screen "Inert Gas Generator Plant" 1280x800, template "Template"
   GraphicView "Graphic view_52" at 522,118 size 43x67; Picture "Graphic_72"
   GraphicView "Graphic view_49" at 715,199 size 43x67; Picture "Graphic_72"
   GraphicView "Graphic view_12" at 522,199 size 43x67; Picture "Graphic_72"
   GraphicView "Graphic view_55" at 522,416 size 43x67; Picture "Graphic_72"
   GraphicView "Graphic view_56" at 650,416 size 43x67; Picture "Graphic_72"
   GraphicView "Graphic view_57" at 522,311 size 43x67; Picture "Graphic_72"
   GraphicView "Graphic view_61" at 527,525 size 32x54; Picture "Graphic_72"
   TextField "Text field_97" at 742,724 size 131x20; Text 'IGG Gas Pressure'
   TextField "Text field_98" at 866,724 size 147x20; Text 'Atom. Air Pressure'
   TextField "Text field_47" at 251,73 size 69x18; Text 'Full Auto'
      Visibility <- "82_To_HMI_CRNT_MODE_IGG"
   TextField "Text field_1" at 251,74 size 55x18; Text 'Manual'
      Visibility <- "82_To_HMI_CRNT_MODE_IGG"
   TextField "Text field_4" at 252,74 size 103x18; Text 'Undetermined'
      Visibility <- "82_To_HMI_CRNT_MODE_IGG"
   TextField "Text field_57" at 252,74 size 36x18; Text 'FAT'
      Visibility <- "82_To_HMI_CRNT_MODE_IGG"
   TextField "Text field_42" at 434,121 size 70x22; Text 'No Flow'
   TextField "Text field_43" at 434,121 size 70x22; Text '- Flow -'
      Visibility <- "10 DI_DATA_FS123"
      Appearance <- "10 DI_DATA_FS123"
   GraphicView "Logo" at 1,1 size 219x60; Picture "Logo of IGG HMI"
   Group "Group_8" at 743,722 size 397x61
   Button "Button_1" at 902,751 size 66x25; TextOn 'Enabled'; TextOff 'Text'
   IOField "I/O field_29" at 898,751 size 70x25; Authorization "Commissioning"; FormatPattern 99.99; Unit  bar
      ProcessValue <- "1111_PID_CV111_Setpoint"
   Group "Group" at 742,724 size 271x20
   IOField "I/O field_10" at 956,109 size 54x22; FormatPattern 999; Unit %
      ProcessValue <- "12_AI_Data_CV403_SCALED"
   IOField "I/O field_15" at 956,95 size 54x22; FormatPattern 999; Unit %
      ProcessValue <- "16_AQ_Data_CV403_CNTRL"
   GraphicView "Graphic view_5" at 1149,212 size 128x29; Picture "Graphic_82"
   GraphicView "Graphic view_91" at 22,264 size 113x127; Picture "Graphic_246"
   GraphicIOField "Graphic I/O field_5" at 14,257 size 129x139; PictureList "New IA Compressor"
      ProcessValue <- "82_To_HMI_IA Compressor Animation"
      Visibility <- "68_Sys_Status_Data_IA_PRES_IN_RNG(1)"
   GraphicView "Graphic view_93" at 147,261 size 48x132; Picture "Graphic_248"
   TextField "Text field_58" at 41,731 size 135x20; Text 'Fuel Pump System'
      Appearance <- "68_Sys_Status_Data_FUEL_PRES_IN_RNG"
   TextField "Text field_89" at 1115,538 size 54x22; Text 'Text'
   Button "HmiScreenItemData_1" at 1,50 size 150x43; TextOn 'Back'; TextOff 'Main Index'
      on Release: ActivateScreen("02 Main Index", 0)
   GraphicView "Graphic view_20" at 336,126 size 900x542; Picture "IGG_5"
   GraphicView "Graphic view_41" at 815,266 size 13x60; Picture "Graphic_57"
   GraphicView "Graphic view_11" at 296,251 size 377x12; Picture "Graphic_20"
   GraphicView "Graphic view_40" at 806,251 size 21x20; Picture "Graphic_41"
   GraphicView "Graphic view_42" at 296,468 size 278x12; Picture "Graphic_20"
   GraphicView "Graphic view_43" at 696,458 size 19x21; Picture "Graphic_40"
   GraphicView "Graphic view_44" at 294,251 size 20x20; Picture "Graphic_42"
   GraphicView "Graphic view_47" at 295,464 size 11x20; Picture "Graphic_56"
   Group "Group_4" at 522,199 size 43x62; Picture "Graphic_72"
   GraphicView "Graphic view_53" at 313,420 size 43x63; Picture "Graphic_72"
   Group "Group_5" at 522,416 size 43x62; Picture "Graphic_72"
   TextField "Text field_2" at 440,182 size 51x16; Text 'FS-123'
   TextField "Text field_3" at 517,182 size 53x16; Text 'CV-124'
   TextField "Text field_5" at 517,263 size 53x16; Text 'CV-215'
   TextField "Text field_7" at 308,375 size 53x16; Text 'CV-111'
   TextField "Text field_8" at 309,479 size 50x16; Text 'CV-203'
   TextField "Text field_9" at 365,479 size 56x16; Text 'PIT-205'
   TextField "Text field_10" at 518,479 size 50x16; Text 'CV-206'
   TextField "Text field_11" at 646,479 size 50x16; Text 'CV-207'
   TextField "Text field_12" at 364,375 size 59x16; Text 'PIT-113'
   TextField "Text field_13" at 441,375 size 48x16; Text 'FS-115'
   TextField "Text field_14" at 517,375 size 53x16; Text 'CV-114'
   GraphicView "Graphic view_15" at 455,338 size 20x26; Picture "Graphic_79"
   GraphicView "Graphic view_16" at 383,339 size 20x26; Picture "Graphic_36"
   GraphicView "Graphic view_51" at 383,444 size 20x26; Picture "Graphic_36"
   TextField "Text field_21" at 80,649 size 55x18; Text 'E-500B'
   GraphicView "Graphic view_2" at 46,502 size 123x15; Picture "Graphic_99"
   GraphicIOField "Graphic I/O field_3" at 75,482 size 60x65; PictureList "Pump Ani"
      ProcessValue <- "82_To_HMI_Fuel Pump 1 Animation"
   GraphicView "Graphic view_6" at 45,604 size 124x15; Picture "Graphic_99"
   GraphicIOField "Graphic I/O field_4" at 75,585 size 60x65; PictureList "Pump Ani"
      ProcessValue <- "82_To_HMI_Fuel Pump 2 Animation"
   GraphicView "Graphic view_8" at 30,517 size 15x94; Picture "Graphic_101"
   GraphicView "Graphic view_9" at 31,593 size 21x25; Picture "Graphic_96"
   GraphicView "Graphic view_10" at 31,503 size 24x23; Picture "Graphic_102"
   GraphicView "Graphic view_25" at 170,517 size 15x94; Picture "Graphic_101"
   GraphicView "Graphic view_26" at 160,503 size 24x23; Picture "Graphic_104"
   GraphicView "Graphic view_29" at 159,594 size 25x24; Picture "Graphic_97"
   GraphicView "Graphic view_30" at 171,553 size 19x24; Picture "Graphic_103"
   GraphicView "Graphic view_33" at 183,557 size 111x15; Picture "Graphic_99"
   GraphicView "Graphic view_48" at 60,502 size 18x15; Picture "Graphic_99"
   GraphicView "Graphic view_58" at 60,604 size 18x15; Picture "Graphic_99"
   TextField "Text field_22" at 80,549 size 56x18; Text 'E-500A'
   GraphicView "Graphic view_76" at 236,534 size 20x26; Picture "Graphic_36"
   IOField "I/O field_1" at 211,512 size 75x18; FormatPattern s99.99; Unit  Bar
      ProcessValue <- "12_AI_Data_PIT204In_SCALED"
   TextField "Text field_23" at 218,576 size 56x16; Text 'PIT-204'
   Rectangle "Rectangle_9" at 66,477 size 78x92
      Appearance <- "10_DI_Data_E500A_TRIPPED"
   Rectangle "Rectangle_10" at 66,580 size 79x92
      Appearance <- "10_DI_Data_E500B_TRIPPED(1)"
   TextField "Text field_24" at 67,673 size 83x18; Text 'Duty Pump'
      Visibility <- "101_Fuel_Pumps_DB_Duty Is B"
   TextField "Text field_25" at 67,457 size 83x18; Text 'Duty Pump'
      Visibility <- "101_Fuel_Pumps_DB_Duty Is A"
   Circle "Circle_11" at 35,559 size 6x6
      Visibility <- "10_DI_Data_E500A_ENBLD"
   GraphicView "Graphic view_46" at 285,547 size 20x24; Picture "Graphic_40"
   GraphicView "Graphic view_21" at 789,331 size 24x10; Picture "Graphic_63"
   GraphicView "Graphic view_22" at 785,326 size 12x13; Picture "Graphic_64"
   GraphicView "Graphic view_23" at 784,176 size 9x156; Picture "Graphic_70"
   GraphicView "Graphic view_27" at 279,176 size 9x185; Picture "Graphic_70"
   GraphicView "Graphic view_35" at 281,363 size 325x11; Picture "Graphic_63"
   GraphicView "Graphic view_39" at 687,379 size 8x10; Picture "Graphic_70"
   GraphicView "Graphic view_38" at 688,386 size 10x13; Picture "Graphic_64"
   GraphicView "Graphic view_7" at 455,147 size 20x26; Picture "Graphic_79"
   GraphicView "Graphic view_18" at 780,172 size 13x15; Picture "Graphic_67"
   GraphicView "Graphic view_14" at 281,171 size 318x11; Picture "Graphic_63"
   GraphicView "Graphic view_17" at 279,172 size 13x15; Picture "Graphic_66"
   Group "Group_2" at 522,118 size 43x62; Picture "Graphic_72"
   GraphicView "Graphic view_31" at 236,331 size 20x26; Picture "Graphic_36"
   IOField "I/O field_6" at 207,308 size 74x18; FormatPattern s99.99; Unit  Bar
      ProcessValue <- "12_AI_Data_PIT112In_SCALED"
   TextField "Text field_17" at 218,375 size 56x16; Text 'PIT-112'
   GraphicView "Graphic view_50" at 313,314 size 43x63; Picture "Graphic_72"
   Group "Group_7" at 522,311 size 43x62; Picture "Graphic_72"
   GraphicView "Graphic view_45" at 293,262 size 13x297; Picture "Graphic_57"
   GraphicView "Graphic view_54" at 305,517 size 24x21; Picture "Graphic_107"
   IOField "I/O field_7" at 358,423 size 77x18; FormatPattern s99.99; Unit  bar
      ProcessValue <- "12_AI_Data_PIT205In_SCALED"
   TextField "Text field_18" at 513,418 size 60x22; Text 'Closed'
      Visibility <- "14_DQ_Data_200CV206ControlOut"
   TextField "Text field_19" at 513,418 size 60x22; Text 'Opened'
      Visibility <- "14_DQ_Data_200CV206ControlOut"
   IOField "I/O field_11" at 330,522 size 55x18; FormatPattern 99.9; Unit  °C
      ProcessValue <- "12_AI_Data_TIT202In_SCALED"
   GraphicView "Graphic view_59" at 558,468 size 145x12; Picture "Graphic_20"
   TextField "Text field_20" at 514,200 size 60x22; Text 'Closed'
   TextField "Text field_26" at 514,200 size 60x22; Text 'Opened'
      Visibility <- "14_DQ_Data_200CV215ControlOut"
   TextField "Text field_31" at 513,315 size 60x22; Text 'Closed'
   TextField "Text field_32" at 513,315 size 60x22; Text 'Opened'
      Visibility <- "14_DQ_Data_200CV114ControlOut"
   TextField "Text field_33" at 305,541 size 56x16; Text 'TIT-202'
   Group "Group_6" at 650,416 size 43x62; Picture "Graphic_72"
   GraphicView "Graphic view_34" at 705,425 size 11x43; Picture "Graphic_57"
   GraphicView "Graphic view_62" at 647,251 size 173x12; Picture "Graphic_20"
   TextField "Text field_28" at 641,419 size 60x22; Text 'Closed'
   TextField "Text field_29" at 641,419 size 60x22; Text 'Opened'
      Visibility <- "14_DQ_Data_200CV207ControlOut"
   GraphicView "Graphic view_63" at 565,171 size 223x11; Picture "Graphic_63"
   Group "Group_3" at 715,199 size 43x62; Picture "Graphic_72"
   TextField "Text field_6" at 710,263 size 53x16; Text 'CV-216'
   TextField "Text field_27" at 706,200 size 60x22; Text 'Closed'
   TextField "Text field_30" at 706,200 size 60x22; Text 'Opened'
      Visibility <- "14_DQ_Data_200CV216ControlOut"
   GraphicView "Graphic view_64" at 581,363 size 107x11; Picture "Graphic_63"
   GraphicView "Graphic view_65" at 695,390 size 12x9; Picture "Graphic_63"
   GraphicView "Graphic view_66" at 851,616 size 24x21; Picture "Graphic_107"
   GraphicView "Graphic view_67" at 1040,616 size 24x21; Picture "Graphic_107"
   IOField "I/O field_8" at 876,617 size 64x18; FormatPattern 99.9; Unit  °C
      ProcessValue <- "12_AI_Data_TIT319_SCALED"
   IOField "I/O field_12" at 1064,617 size 64x18; FormatPattern 99.9; Unit  °C
      ProcessValue <- "12_AI_Data_TIT360_SCALED"
   TextField "Text field_34" at 854,633 size 56x16; Text 'TIT-319'
   TextField "Text field_35" at 1047,633 size 56x16; Text 'TIT-360'
   GraphicView "Graphic view_68" at 1089,539 size 24x21; Picture "Graphic_107"
   TextField "Text field_36" at 1085,559 size 48x16; Text 'LS-001'
   GraphicView "Graphic view_69" at 910,257 size 20x23; Picture "Graphic_36"
   GraphicView "Graphic view_70" at 966,270 size 20x23; Picture "Graphic_36"
   IOField "I/O field_14" at 947,250 size 65x18; FormatPattern s9.99; Unit  bar
      ProcessValue <- "12_AI_Data_PIT316_SCALED"
   GraphicView "Graphic view_71" at 848,241 size 20x26; Picture "Graphic_79"
   TextField "Text field_40" at 433,315 size 70x22; Text 'No Flow'
   TextField "Text field_41" at 433,315 size 70x22; Text '- Flow -'
      Visibility <- "10 DI_DATA_FS115"
      Appearance <- "10 DI_DATA_FS115(1)"
   TextField "Text field_44" at 835,218 size 54x22; Text 'No Flow'
   TextField "Text field_45" at 835,218 size 54x22; Text '- Flow -'
      Visibility <- "10 DI_DATA_FS317"
      Appearance <- "10 DI_DATA_FS317"
   GraphicView "Graphic view_32" at 280,357 size 12x17; Picture "Graphic_64"
   TextField "Text field_48" at 50,404 size 130x20; Text 'I & A Compressor'
      Appearance <- "68_Sys_Status_Data_IA_PRES_IN_RNG"
   GraphicIOField "Graphic I/O field_2" at 273,594 size 196x199; PictureList "IA Compressor_1"
      ProcessValue <- "82_To_HMI_CA Blower Animation"
   GraphicView "Graphic view_13" at 451,640 size 21x27; Picture "Graphic_82"
   GraphicView "Graphic view_36" at 1225,137 size 49x75; Picture "Graphic_108"
   GraphicView "Graphic view_4" at 964,141 size 44x74; Picture "Graphic_108"
   TextField "Text field_50" at 1220,113 size 60x22; Text 'Closed'
      Visibility <- "10_DI_Data_CV401_CLSD"
   IOField "I/O field_5" at 307,295 size 54x22; FormatPattern 999; Unit %
      ProcessValue <- "16_AQ_Data_CV111_CNTRL"
   IOField "I/O field_4" at 307,403 size 54x22; FormatPattern 999; Unit %
      ProcessValue <- "16_AQ_Data_CV203_CNTRL(1)"
   TextField "Text field_52" at 961,125 size 50x16; Text 'CV-403'
   TextField "Text field_53" at 518,576 size 50x16; Text 'CV-127'
   TextField "Text field_56" at 446,576 size 49x16; Text 'PS-101'
   GraphicView "Graphic view_74" at 466,569 size 232x5; Picture "Graphic_63"
   Group "Group_1" at 527,525 size 32x50; Picture "Graphic_72"
   TextField "Text field_54" at 513,526 size 60x22; Text 'Closed'
   TextField "Text field_55" at 513,526 size 60x22; Text 'Opened'
      Visibility <- "14_DQ_Data_200CV127ControlOut"
   GraphicView "Graphic view_73" at 460,550 size 20x26; Picture "Graphic_36"
   GraphicView "Graphic view_75" at 737,434 size 6x141; Picture "Graphic_70"
   GraphicView "Graphic view_78" at 597,569 size 148x5; Picture "Graphic_63"
   GraphicView "Graphic view_3" at 736,566 size 6x8; Picture "Graphic_65"
   GraphicView "Graphic view_28" at 189,356 size 95x11; Picture "Graphic_63"
   GraphicView "Graphic view_19" at 132,317 size 19x12; Picture "Graphic_63"
   GraphicView "Graphic view_72" at 1040,188 size 20x26; Picture "Graphic_36"
   TextField "Text field_59" at 404,73 size 80x18; Text 'Start IGGS'
   TextField "Text field_60" at 340,73 size 70x18; Text 'IA Comp.'
   TextField "Text field_61" at 494,73 size 36x18; Text 'CSW'
   TextField "Text field_62" at 537,73 size 89x18; Text 'Fuel System'
   TextField "Text field_63" at 634,73 size 36x18; Text 'CAB'
   TextField "Text field_64" at 868,72 size 46x18; Text 'Purge'
   TextField "Text field_65" at 806,72 size 52x18; Text 'Pilot B'
   TextField "Text field_66" at 931,72 size 52x18; Text 'Main B'
   TextField "Text field_67" at 1062,72 size 64x18; Text 'Running'
   Circle "Circle_22" at 365,58 size 14x14
      Appearance <- "10 DI_DATA_E131_OK"
   Circle "Circle_23" at 503,58 size 14x14
      Visibility <- "80_From_HMI_RUN_IGG(1)"
      Appearance <- "68_Sys_Status_Data_CSW_IL_PRES_IN_RNG"
   Circle "Circle_24" at 572,58 size 14x14
      Visibility <- "68_Sys_Status_Data_CSW_IL_PRES_IN_RNG"
      Appearance <- "68_Sys_Status_Data_FUEL_PRES_IN_RNG(1)"
   Circle "Circle_25" at 642,58 size 14x14
      Visibility <- "68_Sys_Status_Data_FUEL_PRES_IN_RNG(1)"
      Appearance <- "10_DI_Data_E139_RUNNING"
   Circle "Circle_29" at 1080,55 size 20x20
      Appearance <- "14_DQ_Data_24PF1"
   Circle "Circle_31" at 434,58 size 14x14
      Visibility <- "10 DI_DATA_E131_OK"
      Appearance <- "80_From_HMI_RUN_IGG(1)"
   Circle "Circle_32" at 296,58 size 14x14
      Appearance <- "82_To_HMI_CRNT_MODE_IGG"
   Circle "Circle_27" at 822,58 size 14x14
      Visibility <- "102_Pilot_Burner_DB_FLM_DET"
      Appearance <- "102_Pilot_Burner_DB_RUNNING"
   Circle "Circle_28" at 949,58 size 14x14
      Visibility <- "102_Pilot_Burner_DB_FLM_DET"
      Appearance <- "103_Main_Burner_DB_RUNNING"
   Circle "Circle_9" at 887,58 size 14x14
      Visibility <- "102_Pilot_Burner_DB_FLM_DET"
      Appearance <- "104_Pilot_Purge_DB_DN_OK"
   GraphicView "Graphic view_79" at 132,353 size 19x12; Picture "Graphic_63"
   Button "HmiScreenItemData_9" at 2,97 size 184x29; TextOn 'Back'; TextOff 'IGGS Control'
   Button "HmiScreenItemData_4" at 23,192 size 75x51; TextOn 'Back'; TextOff 'Stop'
      ObjectEnable <- "82_To_HMI_CRNT_MODE_IGG"
      on Release: function_efd93a16("IGG Stop Confirm", 300, 200, -1, -1, 1)
   Circle "Circle_20" at 146,143 size 29x29
      Appearance <- "82_To_HMI_IGG RUN Indication"
   Button "HmiScreenItemData_3" at 23,130 size 75x51; TextOn 'Back'; TextOff 'Start'
      ObjectEnable <- "82_To_HMI_CRNT_MODE_IGG"
      on Release: function_efd93a16("IGG Start Confirm", 300, 200, -1, -1, 1)
   GraphicView "Graphic view_37" at 684,364 size 11x16; Picture "Graphic_67"
   IOField "I/O field_21" at 635,523 size 80x21; FormatPattern s9999; Unit  mBar
      ProcessValue <- "12_AI_Data_PIT102_SCALED(1)"
   TextField "Text field_68" at 644,576 size 56x16; Text 'PIT-102'
   TextField "Text field_15" at 513,121 size 60x22; Text 'Closed'
   TextField "Text field_16" at 513,121 size 60x22; Text 'Opened'
      Visibility <- "14_DQ_Data_200CV124ControlOut"
   Button "HmiScreenItemData_2" at 1128,64 size 150x43; TextOn 'Back'; TextOff 'IGGS Setup'
      on Release: ActivateScreen("Inert Gas Generator Setup", 0)
   GraphicView "Graphic view_77" at 1,556 size 42x15; Picture "Graphic_20"
   GraphicView "Graphic view_85" at 809,353 size 178x145; Picture "Graphic_132"
      Visibility <- "103_Main_Burner_DB_DN_OK(1)"
   GraphicView "Graphic view_82" at 784,321 size 237x221; Picture "Graphic_130"
      Visibility <- "103_Main_Burner_DB_DN_OK(1)"
   GraphicView "Graphic view_86" at 194,566 size 15x144; Picture "Graphic_101"
   GraphicView "Graphic view_87" at 183,704 size 25x21; Picture "Graphic_97"
   TextField "Text field_69" at 1133,358 size 57x18; Text 'Oxygen'
   IOField "I/O field_22" at 1195,354 size 77x27; FormatPattern 99.99; Unit  %
      ProcessValue <- "12_AI_Data_E600O2ContentIn"
   TextField "Text field_70" at 1150,326 size 121x18; Text 'Inert Gas Profile'
   TextField "Text field_71" at 1133,388 size 67x18; Text 'Setpoint'
   TextField "Text field_72" at 1133,426 size 39x18; Text 'Soot'
   IOField "I/O field_24" at 1195,423 size 77x27; FormatPattern 999.9; Unit  %
      ProcessValue <- "12_AI_Data_E700SootContentIn"
   IOField "I/O field_25" at 1195,460 size 77x27; FormatPattern 999.9; Unit  °C
      ProcessValue <- "12_AI_Data_TIT401_SCALED"
   TextField "Text field_73" at 1133,462 size 47x18; Text 'Temp.'
   IOField "I/O field_26" at 1195,496 size 77x27; FormatPattern 9999; Unit  mBar
      ProcessValue <- "12_AI_Data_PIT402_SCALED"
   TextField "Text field_74" at 1133,500 size 65x18; Text 'Pressure'
   GraphicView "Graphic view_89" at 1116,188 size 20x26; Picture "Graphic_36"
   TextField "Text field_39" at 1097,172 size 59x16; Text 'TIT-401'
   IOField "I/O field_18" at 1095,158 size 63x18; FormatPattern 999.9; Unit  °C
      ProcessValue <- "12_AI_Data_TIT401_SCALED"
   TextField "Text field_46" at 446,526 size 50x22; Text 'P'
      Visibility <- "10 DI_DATA_PS101"
   TextField "Text field_75" at 446,526 size 50x22; Text 'No P'
      Visibility <- "10 DI_DATA_PS101"
      Appearance <- "10 DI_DATA_PS101"
   TextField "Text field_77" at 986,271 size 59x16; Text 'PIT-316'
   TextField "Text field_78" at 882,304 size 56x16; Text 'TIT-315'
   TextField "Text field_79" at 793,221 size 48x16; Text 'FS-317'
   IOField "I/O field_3" at 356,319 size 74x18; FormatPattern s99.99; Unit  Bar
      ProcessValue <- "12_AI_Data_PIT113In_SCALED"
   Button "HmiScreenItemData_7" at 215,117 size 150x43; TextOn 'Back'; TextOff 'Air/Fuel Monitoring'
      on Release: ActivateScreen("Air Fuel Monitoring", 0)
   TextField "Text field_51" at 1220,113 size 60x22; Text 'Opened'
      Visibility <- "10_DI_Data_CV401_OPN"
   Button "HmiScreenItemData_11" at 255,608 size 194x179; TextOn 'Back'; TextOff 'Text'
      on Release: ActivateScreen("Air System", 0)
   Line "Line_4" at 812,352 size 3x22
      Visibility <- "14_DQ_Data_X001ControlOut"
   GraphicView "Graphic view_84" at 796,344 size 38x82; Picture "Graphic_129"
      Visibility <- "102_Pilot_Burner_DB_STATE"
   Button "HmiScreenItemData_13" at 741,647 size 358x51; TextOn 'Back'; TextOff 'Cooling System'
      on Release: ActivateScreen("Cooling System", 0)
   IOField "I/O field_23" at 1195,386 size 77x27; Authorization "User administration"; FormatPattern 99.99; Unit  %
      ProcessValue <- "84_Setpoints_E600_BWT_Target"
   TextField "Text field_91" at 465,759 size 169x20; Text 'Combustion Air Blower'
      Appearance <- "10_DI_Data_E139_VSD_FLT"
   TextField "Text field_88" at 835,190 size 54x22; Text 'No Flow'
   TextField "Text field_92" at 835,190 size 54x22; Text '- Flow -'
      Visibility <- "10 DI_DATA_FS320"
      Appearance <- "10 DI_DATA_FS320"
   TextField "Text field_93" at 793,193 size 48x16; Text 'FS-320'
   Button "HmiScreenItemData_18" at 742,647 size 356x51; TextOn 'Back'; TextOff 'Cooling System'
      on Release: ActivateScreen("Cooling System", 0)
      Visibility <- "51_SLAVE_STATUS_P301_ENBLD"
   IOField "I/O field_33" at 462,699 size 72x25; Authorization "Operating Mode"; FormatPattern 9999; Unit  rpm
      ProcessValue <- "80_From_HMI_E139_SET_SPEED"
   IOField "I/O field_34" at 1017,134 size 66x23; FormatPattern 999; Unit  mBar
      ProcessValue <- "19_AUTO_CMNDS_Data_PIT402_Target"
      Appearance <- "19_AUTO_CMNDS_Data_PIT402_Target"
   Button "HmiScreenItemData_19" at 1186,568 size 83x29; TextOn 'Back'; TextOff 'Gas - Trend'
      on Click: function_efd93a16("CV 403 Grafics", 200, 100, -1, -1, 1)
   TextField "Text field_100" at 886,320 size 49x16; Text 'TS-006'
   TextField "Text field_90" at 1117,537 size 54x22; Text 'Text'
   TextField "Text field_38" at 1117,537 size 60x22; Text 'Normal'
      Visibility <- "10 DI_DATA_LS001"
      Appearance <- "10 DI_DATA_LS001"
   TextField "Text field_37" at 1117,537 size 60x22; Text 'Hi Level'
      Visibility <- "10 DI_DATA_LS001"
      Appearance <- "84_Setpoints_TIT315_High"
   GraphicView "Graphic view_90" at 1183,190 size 20x23; Picture "Graphic_36"
   TextField "Text field_103" at 1167,172 size 52x16; Text 'TS-403'
   TextField "Text field_104" at 940,317 size 54x22; Text 'Text'
   TextField "Text field_101" at 940,317 size 54x22; Text 'Hi Temp'
      Visibility <- "10 DI_DATA_TS006(1)"
      Appearance <- "10 DI_DATA_TS006(1)"
   TextField "Text field_102" at 940,317 size 54x22; Text 'Normal'
      Visibility <- "10 DI_DATA_TS006(1)"
   TextField "Text field_107" at 1166,150 size 54x22; Text 'Hi Temp'
      Visibility <- "10 DI_DATA_TS403_FAULT(2)"
      Appearance <- "10 DI_DATA_TS403_FAULT(2)"
   TextField "Text field_108" at 1166,150 size 54x22; Text 'Normal'
      Visibility <- "10 DI_DATA_TS403_FAULT(2)"
      Appearance <- "10 DI_DATA_TS403_FAULT"
   IOField "I/O field_13" at 888,237 size 63x18; FormatPattern 999.9; Unit  °C
      ProcessValue <- "12_AI_Data_TIT315_SCALED"
   IOField "I/O field_20" at 1012,158 size 76x18; FormatPattern s9999; Unit  mBar
      ProcessValue <- "12_AI_Data_PIT402_SCALED"
   GraphicView "Graphic view_88" at 1,713 size 199x13; Picture "Graphic_20"
   TextField "Text field_106" at 886,95 size 59x18; Text 'OPENED'
   GraphicView "Graphic view_1" at 976,199 size 26x62; Picture "Graphic_17"
   TextField "Text field_49" at 1223,246 size 53x16; Text 'CV-401'
   TextField "Text field_76" at 1021,172 size 59x16; Text 'PIT-402'
   GraphicView "Graphic view_60" at 1238,195 size 26x62; Picture "Graphic_17"
   IOField "I/O field_2" at 462,728 size 72x25; FormatPattern 9999; Unit  RPM
      ProcessValue <- "12_AI_Data_E139_RPM_SCALED"
   TextField "Text field_114" at 567,701 size 49x18; Text 'SPEED'
   Button "HmiScreenItemData_15" at 1186,604 size 83x29; TextOn 'Back'; TextOff 'Oxygen'
      on Click: function_efd93a16("CV 203 Grafics", 200, 100, -1, -1, 1)
   IOField "I/O field_28" at 767,752 size 69x23; FormatPattern 999; Unit  mBar
      ProcessValue <- "19_AUTO_CMNDS_Data_PIT402_Target"
      Appearance <- "19_AUTO_CMNDS_Data_PIT402_Target"
   IOField "I/O field_31" at 1034,752 size 80x23; FormatPattern 99.99; Unit  bar
      ProcessValue <- "84_Setpoints_PIT205_Target"
      Appearance <- "84_Setpoints_PIT205_Target"
   TextField "Text field_99" at 1006,724 size 144x20; Text 'Main Fuel Pressure'
   Bar "Bar_1" at 161,270 size 20x105; Unit  %; MinimumValue 0; MaximumValue 100
      ProcessValue <- "12_AI_Data_PIT112In_SCALED"
      MaximumValue <- "84_Setpoints_PIT112_HighHigh"
   TextField "Text field_116" at 52,355 size 57x25; Text 'Enabled'
      Visibility <- "14_DQ_Data_E131ControlOut"
   TextField "Text field_118" at 52,332 size 57x25; Text 'Running'
      Visibility <- "10 DI_DATA_E131_OK"
   Button "HmiScreenItemData_8" at 7,250 size 189x152; TextOn 'Back'; TextOff 'Text'
      on Release: ActivateScreen("Air System", 0)
   IOField "I/O field_17" at 819,414 size 65x25; FormatPattern 999; Unit %
      ProcessValue <- "12_AI_Data_FD001FlameSignalIn"
      Visibility <- "10 DI_DATA_FD001_OK"
   Group "Group_9" at 251,73 size 104x19
   Button "HmiScreenItemData_10" at 14,442 size 178x274; TextOn 'Back'; TextOff 'Text'
      on Release: ActivateScreen("Fuel System", 0)
   DateTimeField "HmiScreenItemData_17" at 1175,0 size 105x30
   DateTimeField "HmiScreenItemData" at 1175,30 size 105x30
   AlarmView "Alarm view_1" at 0,777 size 1280x23
   IOField "I/O field_27" at 744,101 size 83x26; Authorization "Commissioning"; FormatPattern 999; Unit  step
      ProcessValue <- "100_IGG_AUTO_SEQ_DB_CRNT_STEP"
   IOField "I/O field_30" at 744,129 size 83x26; Authorization "Commissioning"; FormatPattern 999; Unit  step
      ProcessValue <- "100_BC_AUTO_SEQ_DB_CRNT_STEP"
   Button "HmiScreenItemData_27" at 633,101 size 83x26; TextOn 'Back'; TextOff 'IGG PLC'
   Button "HmiScreenItemData_28" at 633,129 size 83x26; TextOn 'Back'; TextOff 'BC PLC'
   Group "Group_12" at 677,42 size 115x51
   Circle "Circle_2" at 1013,57 size 14x14
      Visibility <- "102_Pilot_Burner_DB_FLM_DET"
      Appearance <- "19_AUTO_CMNDS_Data_CV203_RAMP_CNTRL"
   TextField "Text field_80" at 984,72 size 82x18; Text 'O2 Control'
   Button "HmiScreenItemData_16" at 209,109 size 376x490; TextOn 'Back'; TextOff 'Text'; Authorization "User administration"
      on Release: ActivateScreen("Air Fuel Monitoring", 0)
   Button "HmiScreenItemData_29" at 770,294 size 329x283; TextOn 'Back'; TextOff 'Text'; Authorization "User administration"
      on Release: ActivateScreen("O2 Content Monitoring", 0)
   Button "HmiScreenItemData_30" at 1098,647 size 176x51; TextOn 'FRESH WATER SYSTEM'; TextOff 'Fresh Water System'; Authorization "Operating Mode"
      on Release: ActivateScreen("Fresh Water System", 0)
      Visibility <- "80_From_HMI_P305_PRSNT"
   Button "HmiScreenItemData_31" at 917,134 size 153x117; TextOn 'Back'; TextOff 'Text'
      on Click: function_efd93a16("CV 403 Grafics", 200, 100, -1, -1, 1)
   GraphicView "Graphic view_81" at 662,544 size 20x26; Picture "Graphic_36"
   Group "Group_10" at 434,121 size 70x22
   GraphicView "Graphic view_83" at 1158,203 size 96x48; Picture "Graphic_235"
   Button "HmiScreenItemData_5" at 1165,191 size 114x70; TextOn 'Back'; TextOff 'Text'
      on Press: ActivateScreen("Inert Gas Conditioning Plant", 0)
   Button "HmiScreenItemData_12" at 1117,260 size 158x52; TextOn 'INERT GAS TRANSFER'; TextOff 'Inert Gas Transfer'; Authorization "Operating Mode"; TextList "IG Transfer"
      on Release: ActivateScreen("IG Transfer Mode", 0)
      ProcessValue <- "80_From_HMI_BWT_BYPASS"
   Button "HmiScreenItemData_14" at 1186,533 size 83x29; TextOn 'Back'; TextOff 'Temp-Trends'
      on Click: function_efd93a16("IGG Temperature Trends", 200, 100, -1, -1, 1)
   Group "Group_11" at 834,364 size 223x284
   Group "Group_13" at 935,209 size 223x226
   Group "Group_14" at 473,288 size 237x372
   Group "Group_15" at 4,254 size 821x468
   Group "Group_16" at 196,173 size 599x224
   GraphicView "Graphic view_24" at 739,597 size 57x58; Picture "Graphic_302"
      Visibility <- "10_DI_Data_IGG_ESTOP_OK"
   Button "HmiScreenItemData_23" at 677,42 size 115x51; TextOn 'Back'; TextOff 'Burner Off'
      Visibility <- "103_Main_Burner_DB_Status"
   Button "HmiScreenItemData_21" at 677,42 size 115x51; TextOn 'Back'; TextOff 'Start Burner'
      Visibility <- "103_Main_Burner_DB_Status"
   Button "HmiScreenItemData_6" at 677,42 size 115x51; TextOn 'Back'; TextOff 'Burner On'
      Visibility <- "103_Main_Burner_DB_Status"
   Button "HmiScreenItemData_22" at 677,42 size 115x51; TextOn 'Back'; TextOff 'Burner Stopped'
      Visibility <- "103_Main_Burner_DB_Status"
   Circle "Circle_104" at 1011,436 size 13x13
      DiagonalMovement <- "CSW_Animation_DB_Animation"
      Visibility <- "10 DI_DATA_FS317"
   Circle "Circle_105" at 1029,410 size 13x13
      DiagonalMovement <- "CSW_Animation_DB_Animation"
      Visibility <- "10 DI_DATA_FS317"
   Circle "Circle_100" at 1038,482 size 13x13
      DiagonalMovement <- "CSW_Animation_DB_Animation"
      Visibility <- "10 DI_DATA_FS317"
   Circle "Circle_98" at 1006,471 size 13x13
      DiagonalMovement <- "CSW_Animation_DB_Animation"
      Visibility <- "10 DI_DATA_FS317"
   Circle "Circle_99" at 1044,458 size 13x13
      DiagonalMovement <- "CSW_Animation_DB_Animation"
      Visibility <- "10 DI_DATA_FS317"
   Circle "Circle_107" at 1038,442 size 13x13
      DiagonalMovement <- "CSW_Animation_DB_Animation"
      Visibility <- "10 DI_DATA_FS317"
   Circle "Circle_94" at 1019,364 size 10x10
      DiagonalMovement <- "CSW_Animation_DB_Animation"
      Visibility <- "10 DI_DATA_FS317"
   Circle "Circle_30" at 1018,602 size 8x8
      Visibility <- "10 DI_DATA_FS317"
      DiagonalMovement <- "CSW_Animation_DB_Animation"
   Circle "Circle_97" at 1028,606 size 8x8
      Visibility <- "10 DI_DATA_FS317"
      DiagonalMovement <- "CSW_Animation_DB_Animation"
   Circle "Circle_102" at 834,640 size 8x8
      DiagonalMovement <- "CSW_Animation_DB_Animation"
      Visibility <- "10 DI_DATA_FS317"
   Circle "Circle_108" at 842,556 size 8x8
      DiagonalMovement <- "CSW_Animation_DB_Animation"
      Visibility <- "10 DI_DATA_FS317"
   Circle "Circle_109" at 953,554 size 8x8
      DiagonalMovement <- "CSW_Animation_DB_Animation"
      Visibility <- "10 DI_DATA_FS317"
   Circle "Circle_96" at 962,520 size 8x8
      DiagonalMovement <- "CSW_Animation_DB_Animation"
      Visibility <- "10 DI_DATA_FS317"
   Circle "Circle_139" at 1074,338 size 10x10
      Visibility <- "51_SLAVE_STATUS_MAIN_BURNER_ACTV"
      VerticalMovement <- "Main Burner Animation_DB_Animation"
   Circle "Circle_134" at 1013,394 size 10x10
      Visibility <- "51_SLAVE_STATUS_MAIN_BURNER_ACTV"
      DiagonalMovement <- "Main Burner Animation_DB_Animation"
   Circle "Circle_135" at 1036,425 size 10x10
      Visibility <- "51_SLAVE_STATUS_MAIN_BURNER_ACTV"
      DiagonalMovement <- "Main Burner Animation_DB_Animation"
   Circle "Circle_136" at 1041,382 size 10x10
      Visibility <- "51_SLAVE_STATUS_MAIN_BURNER_ACTV"
      DiagonalMovement <- "Main Burner Animation_DB_Animation"
   Circle "Circle_137" at 1080,390 size 10x10
      Visibility <- "51_SLAVE_STATUS_MAIN_BURNER_ACTV"
      DiagonalMovement <- "Main Burner Animation_DB_Animation"
   Circle "Circle_143" at 1073,220 size 16x16
      Visibility <- "10_DI_Data_CV401_OPN"
      HorizontalMovement <- "Main Burner Animation_DB_Animation"
   Circle "Circle_144" at 1142,218 size 16x16
      Visibility <- "10_DI_Data_CV401_OPN"
      HorizontalMovement <- "Main Burner Animation_DB_Animation"
   Circle "Circle_146" at 1068,296 size 16x16
      Visibility <- "51_SLAVE_STATUS_MAIN_BURNER_ACTV"
      VerticalMovement <- "Main Burner Animation_DB_Animation"
   Circle "Circle_147" at 1066,217 size 16x16
      Visibility <- "10_DI_Data_CV401_OPN"
      HorizontalMovement <- "Main Burner Animation_DB_Animation"
   Circle "Circle_148" at 1124,217 size 16x16
      Visibility <- "10_DI_Data_CV401_OPN"
      HorizontalMovement <- "Main Burner Animation_DB_Animation"
   Circle "Circle_149" at 1067,277 size 16x16
      Visibility <- "51_SLAVE_STATUS_MAIN_BURNER_ACTV"
      VerticalMovement <- "Main Burner Animation_DB_Animation"
   Circle "Circle_21" at 1069,258 size 10x10
      Visibility <- "51_SLAVE_STATUS_MAIN_BURNER_ACTV"
      VerticalMovement <- "Main Burner Animation_DB_Animation"
   Circle "Circle_145" at 1014,224 size 10x10
      Visibility <- "51_SLAVE_STATUS_MAIN_BURNER_ACTV"
      HorizontalMovement <- "Main Burner Animation_DB_Animation"
   Circle "Circle_150" at 935,209 size 10x10
      Visibility <- "51_SLAVE_STATUS_MAIN_BURNER_ACTV"
      VerticalMovement <- "Main Burner Animation_DB_Animation"
   Circle "Circle_140" at 954,224 size 10x10
      Visibility <- "51_SLAVE_STATUS_MAIN_BURNER_ACTV"
      DiagonalMovement <- "Main Burner Animation_DB_Animation"
   Circle "Circle_133" at 1072,290 size 10x10
      Visibility <- "51_SLAVE_STATUS_MAIN_BURNER_ACTV"
      VerticalMovement <- "Main Burner Animation_DB_Animation"
   Circle "Circle_138" at 1031,354 size 10x10
      Visibility <- "51_SLAVE_STATUS_MAIN_BURNER_ACTV"
      DiagonalMovement <- "Main Burner Animation_DB_Animation"
   Circle "Circle_142" at 1070,424 size 10x10
      Visibility <- "51_SLAVE_STATUS_MAIN_BURNER_ACTV"
      DiagonalMovement <- "Main Burner Animation_DB_Animation"
   Circle "Circle_127" at 473,646 size 14x14
      Visibility <- "10_DI_Data_E139_RUNNING"
      HorizontalMovement <- "82_To_HMI_CA Blower Animation"
   Circle "Circle_126" at 525,646 size 14x14
      Visibility <- "10_DI_Data_E139_RUNNING"
      HorizontalMovement <- "82_To_HMI_CA Blower Animation"
   Circle "Circle_128" at 612,622 size 14x14
      Visibility <- "10_DI_Data_E139_RUNNING"
      VerticalMovement <- "82_To_HMI_CA Blower Animation"
   Circle "Circle_129" at 612,517 size 14x14
      Visibility <- "10_DI_Data_E139_RUNNING"
      VerticalMovement <- "82_To_HMI_CA Blower Animation"
   Circle "Circle_130" at 612,412 size 14x14
      Visibility <- "10_DI_Data_E139_RUNNING"
      VerticalMovement <- "82_To_HMI_CA Blower Animation"
   Circle "Circle_131" at 639,288 size 14x14
      Visibility <- "10_DI_Data_E139_RUNNING"
      HorizontalMovement <- "82_To_HMI_CA Blower Animation"
   Circle "Circle_132" at 696,288 size 14x14
      Visibility <- "10_DI_Data_E139_RUNNING"
      HorizontalMovement <- "82_To_HMI_CA Blower Animation"
   Circle "Circle_26" at 4,561 size 6x6
      Visibility <- "68_Sys_Status_Data_FUEL_PRES_IN_RNG(1)"
      HorizontalMovement <- "Ful Pump Ani Animation_DB_Animation"
   Circle "Circle_3" at 44,508 size 6x6
      Visibility <- "68_Sys_Status_Data_FUEL_PRES_IN_RNG(1)"
      HorizontalMovement <- "IDB_E500A_Animation_Animation"
   Circle "Circle_17" at 43,608 size 6x6
      Visibility <- "68_Sys_Status_Data_FUEL_PRES_IN_RNG(1)"
      HorizontalMovement <- "IDB_E500B_Animation_Animation"
   Circle "Circle_10" at 137,609 size 6x6
      Visibility <- "10_DI_Data_E500B_ENBLD"
      HorizontalMovement <- "IDB_E500B_Animation_Animation"
   Circle "Circle_7" at 134,507 size 6x6
      Visibility <- "10_DI_Data_E500A_ENBLD"
      HorizontalMovement <- "IDB_E500A_Animation_Animation"
   Circle "Circle_19" at 175,517 size 6x6
      Visibility <- "10_DI_Data_E500A_ENBLD"
      VerticalMovement <- "IDB_E500A_Animation_Animation"
   Circle "Circle_18" at 175,596 size 6x6
      Visibility <- "10_DI_Data_E500B_ENBLD"
      VerticalMovement <- "IDB_E500B_Animation_Animation"
   Circle "Circle_35" at 95,716 size 6x6
      Visibility <- "68_Sys_Status_Data_FUEL_PRES_IN_RNG(1)"
      HorizontalMovement <- "Ful Pump Ani Animation_DB_Animation"
   Circle "Circle_51" at 191,716 size 6x6
      Visibility <- "68_Sys_Status_Data_FUEL_PRES_IN_RNG(1)"
      HorizontalMovement <- "Ful Pump Ani Animation_DB_Animation"
   Circle "Circle_52" at 199,643 size 6x6
      Visibility <- "68_Sys_Status_Data_FUEL_PRES_IN_RNG(1)"
      VerticalMovement <- "Ful Pump Ani Animation_DB_Animation"
   Circle "Circle_53" at 199,579 size 6x6
      Visibility <- "68_Sys_Status_Data_FUEL_PRES_IN_RNG(1)"
      VerticalMovement <- "Ful Pump Ani Animation_DB_Animation"
   Circle "Circle_36" at 202,562 size 6x6
      Visibility <- "68_Sys_Status_Data_FUEL_PRES_IN_RNG(1)"
      HorizontalMovement <- "Ful Pump Ani Animation_DB_Animation"
   Circle "Circle_34" at 296,555 size 6x6
      Visibility <- "68_Sys_Status_Data_FUEL_PRES_IN_RNG(1)"
      VerticalMovement <- "Ful Pump Ani Animation_DB_Animation"
   Circle "Circle_49" at 296,456 size 6x6
      Visibility <- "14_DQ_Data_200CV215ControlOut"
      VerticalMovement <- "Ful Pump Ani Animation_DB_Animation"
   Circle "Circle_37" at 307,471 size 6x6
      Visibility <- "14_DQ_Data_200CV206ControlOut"
      HorizontalMovement <- "Ful Pump Ani Animation_DB_Animation"
   Circle "Circle_38" at 402,470 size 6x6
      Visibility <- "14_DQ_Data_200CV206ControlOut"
      HorizontalMovement <- "Ful Pump Ani Animation_DB_Animation"
   Circle "Circle_39" at 498,469 size 6x6
      Visibility <- "14_DQ_Data_200CV206ControlOut"
      HorizontalMovement <- "Ful Pump Ani Animation_DB_Animation"
   Circle "Circle_40" at 593,470 size 6x6
      Visibility <- "14_DQ_Data_200CV206ControlOut"
      HorizontalMovement <- "Ful Pump Ani Animation_DB_Animation"
   Circle "Circle_43" at 707,462 size 6x6
      Visibility <- "14_DQ_Data_200CV207ControlOut"
      VerticalMovement <- "Ful Pump Ani Animation_DB_Animation"
   Circle "Circle_50" at 297,358 size 6x6
      Visibility <- "14_DQ_Data_200CV215ControlOut"
      VerticalMovement <- "Ful Pump Ani Animation_DB_Animation"
   Circle "Circle_48" at 302,254 size 6x6
      Visibility <- "14_DQ_Data_200CV215ControlOut"
      HorizontalMovement <- "Ful Pump Ani Animation_DB_Animation"
   Circle "Circle_47" at 405,254 size 6x6
      Visibility <- "14_DQ_Data_200CV215ControlOut"
      HorizontalMovement <- "Ful Pump Ani Animation_DB_Animation"
   Circle "Circle_46" at 509,254 size 6x6
      Visibility <- "14_DQ_Data_200CV215ControlOut"
      HorizontalMovement <- "Ful Pump Ani Animation_DB_Animation"
   Circle "Circle_45" at 612,254 size 6x6
      Visibility <- "14_DQ_Data_200CV215ControlOut"
      HorizontalMovement <- "Ful Pump Ani Animation_DB_Animation"
   Circle "Circle_44" at 716,254 size 6x6
      Visibility <- "14_DQ_Data_200CV215ControlOut"
      HorizontalMovement <- "Ful Pump Ani Animation_DB_Animation"
   Circle "Circle_42" at 819,282 size 6x6
      Visibility <- "14_DQ_Data_200CV215ControlOut"
      VerticalMovement <- "Ful Pump Ani Animation_DB_Animation"
   Circle "Circle_74" at 196,359 size 6x6
      Visibility <- "68_Sys_Status_Data_IA_PRES_IN_RNG"
      HorizontalMovement <- "IDB_E131_Animation_Animation"
   Circle "Circle_56" at 280,359 size 6x6
      Visibility <- "10 DI_DATA_FS123"
      VerticalMovement <- "IDB_E131_Animation_Animation"
   Circle "Circle_67" at 282,366 size 6x6
      Visibility <- "68_Sys_Status_Data_IA_PRES_IN_RNG"
      HorizontalMovement <- "IDB_E131_Animation_Animation"
   Circle "Circle_68" at 347,366 size 6x6
      Visibility <- "10 DI_DATA_FS115"
      HorizontalMovement <- "IDB_E131_Animation_Animation"
   Circle "Circle_69" at 407,366 size 6x6
      Visibility <- "10 DI_DATA_FS115"
      HorizontalMovement <- "IDB_E131_Animation_Animation"
   Circle "Circle_70" at 473,366 size 6x6
      Visibility <- "10 DI_DATA_FS115"
      HorizontalMovement <- "IDB_E131_Animation_Animation"
   Circle "Circle_71" at 539,366 size 6x6
      Visibility <- "10 DI_DATA_FS115"
      HorizontalMovement <- "IDB_E131_Animation_Animation"
   Circle "Circle_72" at 606,366 size 6x6
      Visibility <- "10 DI_DATA_FS115"
      HorizontalMovement <- "IDB_E131_Animation_Animation"
   Circle "Circle_73" at 690,391 size 6x6
      Visibility <- "10 DI_DATA_FS115"
      HorizontalMovement <- "IDB_E131_Animation_Animation"
   Circle "Circle_64" at 280,281 size 6x6
      Visibility <- "10 DI_DATA_FS123"
      VerticalMovement <- "IDB_E131_Animation_Animation"
   Circle "Circle_57" at 287,174 size 6x6
      Visibility <- "10 DI_DATA_FS123"
      HorizontalMovement <- "IDB_E131_Animation_Animation"
   Circle "Circle_58" at 370,174 size 6x6
      Visibility <- "10 DI_DATA_FS123"
      HorizontalMovement <- "IDB_E131_Animation_Animation"
   Circle "Circle_59" at 453,174 size 6x6
      Visibility <- "10 DI_DATA_FS123"
      HorizontalMovement <- "IDB_E131_Animation_Animation"
   Circle "Circle_60" at 526,174 size 6x6
      Visibility <- "10 DI_DATA_FS123"
      HorizontalMovement <- "IDB_E131_Animation_Animation"
   Circle "Circle_61" at 619,173 size 6x6
      Visibility <- "10 DI_DATA_FS123"
      HorizontalMovement <- "IDB_E131_Animation_Animation"
   Circle "Circle_62" at 703,174 size 6x6
      Visibility <- "10 DI_DATA_FS123"
      HorizontalMovement <- "IDB_E131_Animation_Animation"
   Circle "Circle_65" at 786,179 size 6x6
      Visibility <- "10 DI_DATA_FS123"
      VerticalMovement <- "IDB_E131_Animation_Animation"
   Circle "Circle_66" at 786,262 size 6x6
      Visibility <- "10 DI_DATA_FS123"
      VerticalMovement <- "IDB_E131_Animation_Animation"
   Circle "Circle_63" at 789,333 size 6x6
      Visibility <- "10 DI_DATA_FS123"
      HorizontalMovement <- "IDB_E131_Animation_Animation"

screen "Air Fuel Monitoring" 1280x800, template "Template"
   on GenerateScreen: "TitleUpdater"()
   Gauge "Gauge_1" at 441,189 size 184x184; UnitText '%'; CaptionText 'Open'
      ProcessValue <- "16_AQ_Data_CV111_CNTRL"
   TextField "Text field_10" at 118,229 size 176x20; Text 'Atomising Air Pressure'
   Button "Button_9" at 333,227 size 57x25; TextOn 'Enabled'; TextOff 'Text'
   TextField "Text field_17" at 118,266 size 238x20; Text 'I&A Air Pressure Pilot Setpoint'
   Button "Button_11" at 333,263 size 57x25; TextOn 'Enabled'; TextOff 'Text'
   TextField "Text field_20" at 154,155 size 405x26; Text 'Atomising Air Pressure Control (CV-111)'
   TextField "Text field_12" at 117,339 size 110x20; Text 'Valve Position'
   IOField "I/O field_2" at 333,227 size 74x25; FormatPattern 99.99; Unit  bar
      ProcessValue <- "12_AI_Data_PIT113In_SCALED"
   IOField "I/O field_6" at 333,338 size 74x25; FormatPattern 999.99; Unit  %
      ProcessValue <- "16_AQ_Data_CV111_CNTRL"
   Gauge "Gauge_2" at 441,416 size 184x184; UnitText '%'; CaptionText 'Open'
      ProcessValue <- "16_AQ_Data_CV203_CNTRL(1)"
   TextField "Text field_3" at 118,456 size 160x20; Text 'Burner Fuel Pressure'
   Button "Button_3" at 333,454 size 57x25; TextOn 'Enabled'; TextOff 'Text'
   TextField "Text field_4" at 118,493 size 228x20; Text 'Burner Fuel Pressure Setpoint'
   TextField "Text field_5" at 164,383 size 390x26; Text 'Burner Fuel Pressure Control (CV-203)'
   TextField "Text field_6" at 117,547 size 110x20; Text 'Valve Position'
   IOField "I/O field_1" at 333,454 size 74x25; FormatPattern 99.99; Unit  bar
      ProcessValue <- "12_AI_Data_PIT205In_SCALED"
   IOField "I/O field_5" at 333,546 size 74x25; FormatPattern 999.99; Unit  %
      ProcessValue <- "16_AQ_Data_CV203_CNTRL"
   IOField "I/O field_3" at 333,263 size 74x25; Authorization "Commissioning"; FormatPattern 99.99; Unit  bar
      ProcessValue <- "84_Setpoints_PIT113_Pilot_Target"
   TrendView "Trend view_1" at 703,83 size 572x364
   TrendView "Trend view_2" at 703,475 size 572x255
   Button "HmiScreenItemData_3" at 1,1 size 150x43; TextOn 'Back'; TextOff 'Main Index'
      on Release: ActivateScreen("02 Main Index", 0)
   Button "HmiScreenItemData_1" at 1129,1 size 150x43; TextOn 'I&A Compressor Ok'; TextOff 'Back'
      on Release: function_efd93a16()
   IOField "I/O field_31" at 333,492 size 74x23; FormatPattern 99.99; Unit  bar
      ProcessValue <- "84_Setpoints_PIT205_Target"
      Appearance <- "84_Setpoints_PIT205_Target"
   AlarmView "Alarm view_1" at 0,777 size 1280x23
   Button "HmiScreenItemData_4" at 1129,1 size 150x43; TextOn 'I&A Compressor Ok'; TextOff 'Back'
      on Release: function_efd93a16()
   Group "Group_7" at 213,46 size 373x50
   TextField "Text field_1" at 118,303 size 239x20; Text 'I&A Air Pressure Main Setpoint'
   Button "Button_1" at 333,300 size 57x25; TextOn 'Enabled'; TextOff 'Text'
   IOField "I/O field_4" at 333,300 size 74x25; Authorization "Commissioning"; FormatPattern 99.99; Unit  bar
      ProcessValue <- "84_Setpoints_PIT113_Burner_Target"
   Button "HmiScreenItemData_8" at 227,50 size 355x40; TextOn 'Back'; TextOff 'Text'
   TextField "Screen title" at 213,46 size 373x50; Text 'Screen title'